   REGION "SELECT WIP BUTTON PULSES"
       "Pop Up: Map Select Button Actuations"(screen_elements := #interface.select_wip_buttons,
                                              actuations_as_ints := #actuations_as_ints);
       #"inst WIP Select Button Pulses"(btns := #actuations_as_ints,
                                        pulses := #actuation_pulses_as_ints);
   END_REGION


   REGION "PERFORM WIP SELECTION"
       "Pop Up: Select WIPs: Perform Selection"(indices := #visable_WIPs_indices,
                                                pulses := #actuation_pulses_as_ints,
                                                visable_WIPs:=#visable_WIPs,
                                                selected_wips_as_bools := #t_selected_WIPs_as_Bools);
   END_REGION


   REGION "MAP SELECTION TO META DATA"
       "Pop Up: Select WIPs: Map to Meta"(actuation_pulses_as_ints := #actuation_pulses_as_ints,
                                          indices := #visable_WIPs_indices,
                                          selected_wips_as_bools := #t_selected_WIPs_as_Bools,
                                          selectable_wips := #meta_data.selectable_wips,
                                          selected_wips := #meta_data.selected_wips);
   END_REGION    


   REGION "HOUSE KEEPING FOR STATION SELECTION CHANGE"
       IF #meta_data.selection_change.selection_change THEN
           "Array.DInt.Fill"(int_in := INT_TO_DINT("NULL_TOKEN"),
                             array_out => #visable_WIPs);
           FOR #i := 0 TO "WIP_COUNT" DO
               #t_selected_WIPs_as_Bools[#i] := FALSE;
           END_FOR;
           "Clear WIP Selection Meta Data"(#meta_data.selected_wips);
       END_IF;
   END_REGION


   REGION "BUILD SELECTABLE WIP LIST"
       IF #meta_data.selection_change.selection_change THEN
           IF "Is_HMI_Station"(#stations.stn[#meta_data.selection_change.station_index]) THEN
               "Pop Up: Select WIPs: Build Selectable List"(saved_WIPs := #saved_WIPs,
                                                            meta_data := #meta_data,
                                                            stations := #stations);
           END_IF;
       END_IF;
   END_REGION


   REGION "SHOW ALL WIPS WHEN FEWER SELECTABLE WIPS THAN BUTTONS"
       IF #meta_data.selection_change.selection_change AND #meta_data.selectable_wips.count - 1 <= "WIP_POPUP_BUTTON_COUNT" THEN
           "Array.DInt.Fill"(int_in := INT_TO_DINT("NULL_TOKEN"),
                             array_out => #visable_WIPs_indices);
           FOR #i := 0 TO #meta_data.selectable_wips.count - 1 DO
               #visable_WIPs[#i] := #meta_data.selectable_wips.wips[#i];
               #visable_WIPs_indices[#i] := #i;
           END_FOR;
       END_IF;
   END_REGION



   REGION "NAVIGATE THROUGH TABLE WHEN MORE SELECTABLE WIPS THAN BUTTONS"
       IF #meta_data.selectable_wips.count - 1 > "WIP_POPUP_BUTTON_COUNT" THEN

           REGION "TABLE NAVIGATION"
               #"inst Table Nav"(first_null_index := #meta_data.selectable_wips.count,
                                 tblData := #meta_data.selectable_wips.wips,
                                 tblDisp := #visable_WIPs,
                                 tableNav := #interface.nav_bar.plc,
                                 rowIndices := #visable_WIPs_indices);
           END_REGION

           REGION "MAP INDICES ON SCANS WHEN SELECTION HASN'T CHANGED"
               IF NOT #meta_data.selection_change.selection_change THEN
                   FOR #i := 0 TO "WIP_POPUP_BUTTON_COUNT" DO
                       #visable_WIPs[#i] := #meta_data.selectable_wips.wips[#visable_WIPs_indices[#i]];
                   END_FOR;
               END_IF;
           END_REGION

           REGION "REMAP INDICES TO TOP WHEN SELECTION HAS CHANGED"
               IF #meta_data.selection_change.selection_change THEN
                   FOR #i := 0 TO "WIP_POPUP_BUTTON_COUNT" DO
                       #visable_WIPs[#i] := INT_TO_DINT(#i);
                       #visable_WIPs_indices[#i] := INT_TO_DINT(#i);
                   END_FOR;
               END_IF;
           END_REGION

       END_IF;
   END_REGION
END_FUNCTION_BLOCK

FUNCTION "Pop Up: Select WIPs: Get Matching WIPs" : Void   // FC125, SCL
{ S7_Optimized_Access := 'TRUE' }
VERSION : 0.1
   VAR_INPUT
      selectable_wips : "Selectable Wips";
      station_wips : "Selectable Wips";
   END_VAR
   VAR_IN_OUT
      matching_wips : "Selectable Wips";
   END_VAR
   VAR_TEMP
      i : Int;
      j : Int;
      t_matching_wips : "Selectable Wips";
   END_VAR
BEGIN
   REGION "COPY TO LOCAL"
       "Array.DInt.Fill"(int_in := INT_TO_DINT("NULL_TOKEN"),
                         array_out => #t_matching_wips.wips);
       #t_matching_wips.count := 0;
   END_REGION

   REGION "COMPARE EACH WIP CODE IN OUTER LIST ..." 
       FOR #i := 0 TO "WIP_COUNT" DO

           REGION "LEAVE LOOP ON FIRST NULL"
               IF #selectable_wips.wips[#i] = "NULL_TOKEN" THEN
                   EXIT;
               END_IF;
           END_REGION

           REGION "WITH EACH IN INNER LIST AND ..."
               FOR #j := 0 TO "WIP_COUNT" DO

                   REGION "LEAVE LOOP ON FIRST NULL"
                       IF #station_wips.wips[#j] = "NULL_TOKEN" THEN
                           EXIT;
                       END_IF;
                   END_REGION

                   REGION "COPY MATCHES"
                       IF #selectable_wips.wips[#i] = #station_wips.wips[#j] THEN
                           #t_matching_wips.wips[#t_matching_wips.count] := #selectable_wips.wips[#i];
                           #t_matching_wips.count += 1;
                       END_IF;
                   END_REGION

               END_FOR;
           END_REGION

       END_FOR;
   END_REGION


   REGION "RETURN"
       #matching_wips := #t_matching_wips;
   END_REGION
END_FUNCTION

FUNCTION "Pop Up: Select WIPs: Build Selectable List" : Void   // FC128, SCL
{ S7_Optimized_Access := 'TRUE' }
VERSION : 0.1
   VAR_INPUT
      stations : "Station: All Stations";
      saved_WIPs : "Recipe: HMI Stations Saved Wips";
   END_VAR
   VAR_IN_OUT
      meta_data : "Setting Meta Data";
   END_VAR
   VAR_TEMP
      wip_index : Int;
      p_outer : Int;
      p_inner : Int;
      t_selectable_WIPs : "Selectable Wips";
      selected_station_WIPs : "Selected Wips";
   END_VAR
BEGIN
   REGION "NO STATIONS SELECTED"
       IF #meta_data.selected_stations.count = 0 THEN
           "Array.DInt.Fill"(int_in := INT_TO_DINT("NULL_TOKEN"),
                             array_out => #t_selectable_WIPs.wips);
           #t_selectable_WIPs.count := 0;
           GOTO RTRN;
       END_IF;
   END_REGION


   REGION "SINGLE STATION SELECTION"
       IF #meta_data.selected_stations.count = 1 THEN
           "Array.DInt.Fill"(int_in := -1,
                             array_out => #t_selectable_WIPs.wips);
           #t_selectable_WIPs.count := 0;
           #wip_index := "WIP.Global_Index_to_HMI_Station_Index"(global_index := "Get First Selected Station"(#meta_data.selected_stations.stns),
                                                                 saved_WIPs := #saved_WIPs);
           "Pop Up: Select WIPs: Map WIP Codes"(wip_station := #saved_WIPs.stn[#wip_index],
                                                selectable_wips := #t_selectable_WIPs);
           GOTO RTRN;
       END_IF;
   END_REGION


   REGION "MULTI STATION SELECTION"

       REGION "CHECK MATCHING: SELECTABLE & NEW STATION"
           #t_selectable_WIPs.wips := #meta_data.selectable_wips.wips;
           "Array.DInt.Fill"(int_in := INT_TO_DINT("NULL_TOKEN"),
                             array_out => #selected_station_WIPs.wips);
           "Map WIP Codes to DInt Array"(station := "WIP.Global_Index_to_Station"(index := #meta_data.selection_change.station_index, wip_stations := #saved_WIPs),
                                         WIP_array := #selected_station_WIPs.wips);
           "Pop Up: Select WIPs: Get Matching WIPs"(selectable_wips := #meta_data.selectable_wips,
                                                    station_wips := #selected_station_WIPs,
                                                    matching_wips := #t_selectable_WIPs);
       END_REGION


   END_REGION


   REGION "RETURN"
   RTRN:
       #meta_data.selectable_wips := #t_selectable_WIPs;
   END_REGION
END_FUNCTION

FUNCTION "Pop Up: Select WIPs: Map WIP Codes" : Void   // FC129, SCL
{ S7_Optimized_Access := 'TRUE' }
VERSION : 0.1
   VAR_INPUT
      wip_station : "WIP: Station";
   END_VAR
   VAR_IN_OUT
      selectable_wips : "Selectable Wips";
   END_VAR
   VAR_TEMP
      i : Int;
      t_selectable_wips : "Selectable Wips";
   END_VAR
BEGIN
   REGION "COPY TO LOCAL"
       #t_selectable_wips := #selectable_wips;
   END_REGION


   REGION "MAP VALUES"
       "Map WIP Codes to DInt Array"(station := #wip_station,
                                     WIP_array := #t_selectable_wips.wips);
   END_REGION


   REGION "COUNT SELECTABLE WIPS"
       #t_selectable_wips.count := "Count Collapsed DInt Array"(null_value := INT_TO_DINT("NULL_TOKEN"),
                                                                array := #t_selectable_wips.wips);
   END_REGION


   REGION "RETURN"
       #selectable_wips := #t_selectable_wips;
   END_REGION
END_FUNCTION

FUNCTION "Pop Up: Select WIPs: Animations" : Void   // FC134, SCL
{ S7_Optimized_Access := 'TRUE' }
VERSION : 0.1
   VAR_INPUT
      selectable_WIP_count : Int;
      selected_WIPs : Array[0.."WIP_COUNT"] of Bool;
      visable_WIPs : Array[0.."WIP_POPUP_BUTTON_COUNT"] of DInt;
      visable_WIPs_indices : Array[0.."WIP_POPUP_BUTTON_COUNT"] of Int;
      wip_library : "Recipe: Wip Text Library";
   END_VAR
   VAR_IN_OUT
      interface : "Select WIP";
   END_VAR
   VAR_TEMP
      i : Int;
      labels : Array[0.."WIP_POPUP_BUTTON_COUNT"] of String;
      t_interface : "Select WIP";
      t_selected_WIPs : Array[0.."WIP_COUNT"] of Int;
      visable_WIP_count : Int;
   END_VAR
BEGIN
   REGION "COPY TO LOCAL"
       #t_interface := #interface;
   END_REGION


   REGION "ANIMATE CLOSE SCREEN BUTTON"
       #t_interface.close_screen.animate := "Bool.Animate"(true_color := "GREEN_LIGHT_BACKGROUND",
                                                           false_color := "RED_LIGHT_BACKGROUND",
                                                           evaluation_signal := #t_interface.close_screen.actuate);
   END_REGION


   REGION "ANIMATE WIP SELECT BUTTONS" 

       REGION "WIP LABELS"
           FOR #i := 0 TO "WIP_POPUP_BUTTON_COUNT" DO
               #labels[#i] := WSTRING_TO_STRING("WIP.Code_to_WString"(wipTxtLib := #wip_library, code := #visable_WIPs[#i]));
           END_FOR;
       END_REGION

       REGION "CONVERT BOOLS TO INT FOR MOVE BLOCK VARIANT"
           FOR #i := 0 TO "WIP_COUNT" DO
               #t_selected_WIPs[#i].%X0 := #selected_WIPs[#i];
           END_FOR;
       END_REGION

       REGION "ANIMATE"
           #visable_WIP_count := "Count Collapsed DInt Array"(null_value := INT_TO_DINT("NULL_TOKEN"),
                                                              array := #visable_WIPs);
           "Animate Array: PB Data"(labels := #labels,
                                    pb_data := #t_interface.select_wip_buttons,
                                    selected_elements := #t_selected_WIPs,
                                    visible_elements := #visable_WIPs_indices,
                                    visible_pb_count := #visable_WIP_count);
       END_REGION

   END_REGION


   REGION "NAV BAR"
       "Pop Up: Nav Bar: Animate"(selectable_element_count := #selectable_WIP_count - 1,
                                  visible_rows := "WIP_POPUP_BUTTON_COUNT",
                                  nav_bar := #t_interface.nav_bar);
   END_REGION


   REGION "DRAW"
       #interface := #t_interface;
   END_REGION
END_FUNCTION

FUNCTION "Pop Up: Select WIPs: Perform Selection" : Void   // FC137, SCL
{ S7_Optimized_Access := 'TRUE' }
VERSION : 0.1
   VAR_INPUT
      indices : Array[0.."WIP_POPUP_BUTTON_COUNT"] of DInt;
      pulses : Array[0.."WIP_POPUP_BUTTON_COUNT"] of Int;
      visable_WIPs : Array[0.."WIP_POPUP_BUTTON_COUNT"] of DInt;
   END_VAR
   VAR_IN_OUT
      selected_wips_as_bools : Array[0.."WIP_COUNT"] of Bool;
   END_VAR
   VAR_TEMP
      i : Int;
      t_selected_wips_as_bools : Array[0.."WIP_COUNT"] of Bool;
   END_VAR
BEGIN
   REGION "NOTES"
       (*
           The same wip code can exist in several hmi stations, so 
           selected wips are stored by generating an array of codes.
           Later, the codes can be checked at each station for station 
           modificatins.
           This function starts the process by checking the visable indices
           array (a list of pointers to rows in the selectable wip array).
           If an actuation occurs on a button, visible[x] will give the row 
           number of the wip code in the selectable wip array.
           The row number in the selected wip array is then set to true.
           The toggeled state together with the pulse allows the selected 
           wips list to be rebuilt easily.
       *)
   END_REGION


   REGION "COPY TO LOCAL"
       #t_selected_wips_as_bools := #selected_wips_as_bools;
   END_REGION


   REGION "CHECK INDEX ARRAY"
       FOR #i := 0 TO "WIP_POPUP_BUTTON_COUNT" DO

           REGION "EXIT ON NULL"
               IF #visable_WIPs[#i] = "NULL_TOKEN" THEN
                   EXIT;
               END_IF;
           END_REGION

           REGION "TOGGLE WIP SELECT STATE"
               "Toggle"(pulse := #pulses[#i].%X0,
                        state := #t_selected_wips_as_bools[DINT_TO_INT(#indices[#i])]);
           END_REGION

       END_FOR;
   END_REGION


   REGION "RETURN"
       #selected_wips_as_bools := #t_selected_wips_as_bools;
   END_REGION
END_FUNCTION

FUNCTION "Pop Up: Select WIPs: Map to Meta" : Void   // FC138, SCL
{ S7_Optimized_Access := 'TRUE' }
VERSION : 0.1
   VAR_INPUT
      actuation_pulses_as_ints : Array[0.."WIP_POPUP_BUTTON_COUNT"] of Int;
      indices : Array[0.."WIP_POPUP_BUTTON_COUNT"] of DInt;
      selected_wips_as_bools : Array[0.."WIP_COUNT"] of Bool;
      selectable_wips : "Selectable Wips";
   END_VAR
   VAR_IN_OUT
      selected_wips : "Selected Wips";
   END_VAR
   VAR_TEMP
      rebuild_selected_wips : Bool;
      i : Int;
      t_selected_wips : "Selected Wips";
   END_VAR
BEGIN
   REGION "NOTES"
       (*
           This function has two states.
           The first state checks for any selection pulse.
           On such a pulse, the selected wip code array is filled
           with nulls, the selected wip counter is reset, and the 
           state flag to rebuild the array is set.
           In the rebuild array state, each element of the selected
           wip array of bools is checked. 
           If true, the code from the corresponding selectable wip
           code array is saved to the selected wip code array and 
           the selected wip count is incremented.
           When this function has completed, the array of selected wips
           in meta data section of the hmi settings db will be up to 
           date.
          *)
   END_REGION


   REGION "COPY TO LOCAL"
       #t_selected_wips := #selected_wips;
   END_REGION


   REGION "SCAN FOR PULSES, INITIALIZE AND SET STATE"
       FOR #i := 0 TO "WIP_POPUP_BUTTON_COUNT" DO
           IF #actuation_pulses_as_ints[#i].%X0 THEN
               "Array.DInt.Fill"(int_in := INT_TO_DINT("NULL_TOKEN"),
                                 array_out => #t_selected_wips.wips);
               #t_selected_wips.count := 0;
               #rebuild_selected_wips := TRUE;
               EXIT;
           END_IF;
       END_FOR;
   END_REGION


   REGION "REBUILD ARRAY, INCREMENT SELECTED WIP COUNT"
       IF #rebuild_selected_wips THEN
           FOR #i := 0 TO "WIP_COUNT" DO
               IF #selected_wips_as_bools[#i] THEN
                   #t_selected_wips.wips[#t_selected_wips.count] := #selectable_wips.wips[#i];
                   #t_selected_wips.count += 1;
               END_IF;
           END_FOR;
       END_IF;
   END_REGION


   REGION "RETURN"
       #selected_wips := #t_selected_wips;
   END_REGION
END_FUNCTION

// folder: HMI: Warehouse/RSP Simulation

FUNCTION_BLOCK "Sim: from Global"   // FB26, SCL
{ S7_Optimized_Access := 'TRUE' }
VERSION : 0.1
   VAR_INPUT
      stns : "Station: All Stations";
   END_VAR
   VAR_IN_OUT
      simStations : "Simulated Stations";
   END_VAR
   VAR
      old : Struct
         nextGrp : Bool;
         prevGrp : Bool;
      END_STRUCT;
   END_VAR
   VAR_TEMP
      animate : USInt;
      btnCount : Int;
      currentBtn : Bool;
      dzLabel : WString;
      firstStn : Int;
      i : Int;
      intBox : Int;
      j : Int;
      kp8Color : DWord;
      label : WString;
      oldBtn : Bool;
      pSim : Int;
      pStn : Int;
   END_VAR
   VAR CONSTANT
      space : WString := WSTRING#' ';
      lead0 : WString := WSTRING#'0';
      volvo16 : WString := WSTRING#'VOLVO 16';
   END_VAR
BEGIN
   REGION "COPY TO LOCAL"
       #firstStn := #simStations.firstStn;
   END_REGION

   REGION "RESOLVE STATION POINTER"

       REGION "PROCESS NEXT GROUP PRESS"

           REGION "COPY TO LOCAL"
               #currentBtn := #simStations.down.actuate;
               #oldBtn := #old.nextGrp;
           END_REGION

           REGION "FALLING EDGE OF NEXT GROUP"
               IF NOT #currentBtn AND #oldBtn THEN

                   REGION "INCREMENT FIRST STATION"
                       #firstStn += "simKP8Count";
                   END_REGION

                   REGION "UPPER LIMIT ROLL OVER"
                       IF #firstStn > "STATION_COUNT" THEN
                           #firstStn -= "STATION_COUNT" + 1;
                       END_IF;
                   END_REGION

               END_IF;
           END_REGION

           REGION "NEXT GROUP CHANGE DETECTION"
               #old.nextGrp := #currentBtn;
           END_REGION

       END_REGION

       REGION "PROCESS PREVIOUS GROUP PRESS"

           REGION "COPY TO LOCAL"
               #currentBtn := #simStations.up.actuate;
               #oldBtn := #old.prevGrp;
           END_REGION

           REGION "FALLING EDGE OF PREVIOUS GROUP"
               IF NOT #currentBtn AND #oldBtn THEN

                   REGION "DECREMENT FIRST STATION"
                       #firstStn -= "simKP8Count";
                   END_REGION

                   REGION "LOWER LIMIT ROLL OVER"
                       IF #firstStn < 0 THEN
                           #firstStn += "STATION_COUNT" + 1;
                       END_IF;
                   END_REGION

               END_IF;
           END_REGION

           REGION "PREVIOUS GROUP CHANGE DETECTION"
               #old.prevGrp := #currentBtn;
           END_REGION

       END_REGION

   END_REGION

   REGION "FOR EACH BUTTON"
       FOR #i := 0 TO 11 DO

           REGION "CALCULATE POINTER"
               #pStn := #i + #firstStn;
               #pSim := #i;
           END_REGION

           REGION "UPPER LIMIT ROLL OVER"
               IF #pStn > "STATION_COUNT" THEN
                   #pStn := #firstStn + #i - "STATION_COUNT" - 1;
               END_IF;
           END_REGION

           REGION "COPY TO LOCAL"
               #kp8Color := #stns.stn[#pStn].wipCmpts.ioData.kp8.tempOut;
           END_REGION

           REGION "LABEL STATIONS"

               REGION "DETERMINE LINE LABEL"
                   #label := #stns.stn[#pStn].id.lineName;
                   IF #label = #volvo16 THEN
                       #label := WSTRING#'V16';
                   END_IF;
               END_REGION

               REGION "DETERMINE DROP ZONE LABEL"
                   #intBox := USINT_TO_INT(#stns.stn[#pStn].id.dropZone);
                   IF #intBox <= 9 THEN
                       #dzLabel := CONCAT_WSTRING(IN1 := #lead0,
                                                  IN2 := "Strip Sign"(INT_TO_WSTRING(#intBox)));
                   END_IF;
                   IF #intBox >= 10 THEN
                       #dzLabel := "Strip Sign"(INT_TO_WSTRING(#intBox));
                   END_IF;
               END_REGION

               REGION "WRITE LABEL"
                   #label := CONCAT_WSTRING(IN1 := #label,
                                            IN2 := #space,
                                            IN3 := #dzLabel);
                   #simStations.me[#pSim].stn.label := #label;
               END_REGION

           END_REGION

           REGION "ANIMATE STATION LABEL"
               #simStations.me[#pSim].stn.animate := "GRAY_BACKGROUND";
           END_REGION

           REGION "FOR EACH BUTTON"
               FOR #j := 0 TO "STATION_BUTTON_COUNT" DO

                   REGION "COLOR BUTTONS"
                       #animate := "KP8 Driver: HMI Emulator: Animation"(kp8Color := #kp8Color,
                                                                btnNumber := #j);
                       #simStations.me[#pSim].btn.animate[#j] := #animate;
                   END_REGION

                   REGION "WRITE BUTTON LABELS"
                       #intBox := "Pointer Calc: KP8 Labels"(#j);
                       #label := "Strip Sign"(INT_TO_WSTRING(#intBox));
                       #simStations.me[#pSim].btn.labels[#j] := #label;
                   END_REGION

               END_FOR;
           END_REGION

       END_FOR;
   END_REGION

   REGION "SAVE FIRST STATION"
       #simStations.firstStn := #firstStn;
   END_REGION

   REGION "ANIMATE NEXT GROUP PRESS"
       #simStations.down.animate := "Bool.Animate"(true_color := "GREEN_LIGHT_BACKGROUND",
                                                   false_color := "GRAY_BACKGROUND",
                                                   evaluation_signal := #simStations.down.actuate);
   END_REGION

   REGION "ANIMATE PREV GROUP PARESS"
       #simStations.up.animate := "Bool.Animate"(true_color := "GREEN_LIGHT_BACKGROUND",
                                                 false_color := "GRAY_BACKGROUND",
                                                 evaluation_signal := #simStations.up.actuate);
   END_REGION
END_FUNCTION_BLOCK

FUNCTION "Sim: to Global" : Void   // FC23, SCL
{ S7_Optimized_Access := 'TRUE' }
VERSION : 0.1
   VAR_INPUT
      simStns : "Simulated Stations";
   END_VAR
   VAR_IN_OUT
      stations : "Station: All Stations";
   END_VAR
   VAR_TEMP
      i : Int;
      j : Int;
      pSim : Int;
      pStn : Int;
   END_VAR
BEGIN
   REGION "COPY TO LOCAL"
       // #btnCount := "btnCount";
       // #firstStn := #simStns.firstStn;
       // #simKP8Count := "simKP8Count";
       // #stnCount := "stnCount";
   END_REGION

   REGION "FOR EACH STATION"
       FOR #i := 0 TO "simKP8Count" DO

           REGION "CALCULATE POINTER"
               #pStn := #i + #simStns.firstStn;
               #pSim := #i;
           END_REGION

           REGION "UPPER LIMIT ROLL OVER"
               IF #pStn > "STATION_COUNT" THEN
                   #pStn := #simStns.firstStn + #i - "STATION_COUNT" - 1;
               END_IF;
           END_REGION

           REGION "COPY SIMULATED PRESSES"
               #stations.stn[#pStn].wipCmpts.ioData.kp8.input.%B1 := #simStns.me[#pSim].btn.actuate;
           END_REGION

       END_FOR;
   END_REGION
END_FUNCTION

FUNCTION "Sim: KP8 Animations" : Word   // FC84, SCL
{ S7_Optimized_Access := 'TRUE' }
VERSION : 0.1
   VAR_INPUT
      pbs : DWord;
   END_VAR
   VAR_TEMP
      ret : Word;
   END_VAR
BEGIN
   #"Sim: KP8 Animations".%B1 := #pbs.%B0;
   #"Sim: KP8 Animations".%B0 := #pbs.%B1;
END_FUNCTION

// folder: Linked List

FUNCTION_BLOCK "Linked List"   // FB29, SCL
{ S7_Optimized_Access := 'TRUE' }
VERSION : 0.1
   VAR_IN_OUT
      interface : "Linked List: Method Interface";
   END_VAR
   VAR
      list : "Linked List: List";
   END_VAR
   VAR CONSTANT
      TERMINAL_BEHAVIOR : String := 'open';
   END_VAR
BEGIN
   REGION "APPEND"
       IF #interface.append.in.request THEN
           "Linked List: Append"(terminal_behavior := #TERMINAL_BEHAVIOR,
                                 commands := #interface.append,
                                 list := #list);
       END_IF;
   END_REGION

   REGION "DELETE"
       IF #interface.delete.in.request THEN
           "Linked List: Delete"(commands := #interface.delete,
                                 list := #list);
       END_IF;
   END_REGION

   REGION "DISPLAY"
       IF #interface.display.in.request THEN
           "Linked List: Display"(commands := #interface.display,
                                  list := #list);
       END_IF;
   END_REGION

   REGION "INSERT"
       IF #interface.insert.in.request THEN
           "Linked List: Insert"(terminal_behavior := #TERMINAL_BEHAVIOR,
                                 commands := #interface.insert,
                                 list := #list);
       END_IF;
   END_REGION

   REGION "RESET"
       IF #interface.reset.in.request THEN
           "Linked List: Reset"(commands := #interface.reset,
                                list := #list);
       END_IF;
   END_REGION

   REGION "REVERSE"
       IF #interface.reverse.in.request THEN
           "Linked List: Reverse"(commands := #interface.reverse,
                                  list := #list);
       END_IF;
   END_REGION

   REGION "SEARCH"
       IF #interface.search.in.request THEN
           "Linked List: Search"(commands := #interface.search,
                                 list := #list);
       END_IF;
   END_REGION
END_FUNCTION_BLOCK

FUNCTION "Linked List: Private: Clear Node" : Void   // FC156, SCL
{ S7_Optimized_Access := 'TRUE' }
VERSION : 0.1
   VAR_IN_OUT
      node : "Linked List: Node";
   END_VAR
   VAR_TEMP
      ret : "Linked List: Node";
   END_VAR
BEGIN
   #ret.meta.key := "NULL_TOKEN";
   #ret.meta.next := "NULL_TOKEN";
   #node := #ret;
END_FUNCTION

FUNCTION "Linked List: Private: Get Head" : "Linked List: Node"   // FC157, SCL
{ S7_Optimized_Access := 'TRUE' }
VERSION : 0.1
   VAR_INPUT
      list : "Linked List: List";
   END_VAR
   VAR_TEMP
      pointer_list : DInt;
      ret : "Linked List: Node";
   END_VAR
BEGIN
   FOR #pointer_list := 0 TO "LINKED_LIST_LENGTH" DO
       IF #list.me[#pointer_list].meta.is_head THEN
           #ret := #list.me[#pointer_list];
           EXIT;
       END_IF;
   END_FOR;
   #"Linked List: Private: Get Head" := #ret;
END_FUNCTION

FUNCTION "Linked List: Private: Before" : Void   // FC158, SCL
{ S7_Optimized_Access := 'TRUE' }
VERSION : 0.1
   VAR_IN_OUT
      next_node : "Linked List: Node";   // next_node goes after node
      node : "Linked List: Node";   // node goes before next_node
   END_VAR
BEGIN
   #node.meta.next := #next_node.meta.key;
   IF #next_node.meta.is_head THEN
       #next_node.meta.is_head := FALSE;
       #node.meta.is_head := TRUE;
   END_IF;
END_FUNCTION

FUNCTION "Linked List: Private: Tail Swap" : Void   // FC159, SCL
{ S7_Optimized_Access := 'TRUE' }
VERSION : 0.1
   VAR_IN_OUT
      new_tail : "Linked List: Node";
      old_tail : "Linked List: Node";
   END_VAR
BEGIN
   #new_tail.meta.is_tail := TRUE;
   #old_tail.meta.is_tail := FALSE;
END_FUNCTION

FUNCTION "Linked List: Private: Head Swap" : Void   // FC160, SCL
{ S7_Optimized_Access := 'TRUE' }
VERSION : 0.1
   VAR_IN_OUT
      new_head : "Linked List: Node";
      old_head : "Linked List: Node";
   END_VAR
BEGIN
   #new_head.meta.is_head := TRUE;
   #old_head.meta.is_head := FALSE;
END_FUNCTION

FUNCTION "Linked List: Private: Get Next" : "Linked List: Node"   // FC161, SCL
{ S7_Optimized_Access := 'TRUE' }
VERSION : 0.1
   VAR_INPUT
      current : "Linked List: Node";
      list : "Linked List: List";
   END_VAR
   VAR_TEMP
      ret : "Linked List: Node";
   END_VAR
BEGIN
   "Linked List: Private: Clear Node"(#ret);
   IF #list.me[#current.meta.key].meta.next <> "NULL_TOKEN" THEN
       #ret := #list.me[#current.meta.next];
   END_IF;
   #"Linked List: Private: Get Next" := #ret;
END_FUNCTION

FUNCTION "Linked List: Private: Get Previous" : "Linked List: Node"   // FC162, SCL
{ S7_Optimized_Access := 'TRUE' }
VERSION : 0.1
   VAR_INPUT
      current : "Linked List: Node";
      list : "Linked List: List";
   END_VAR
   VAR_TEMP
      list_pointer : DInt;
      ret : "Linked List: Node";
   END_VAR
BEGIN
   "Linked List: Private: Clear Node"(#ret);
   FOR #list_pointer := 0 TO "LINKED_LIST_LENGTH" DO
       IF #list.me[#list_pointer].meta.next = #current.meta.key THEN
           #ret := #list.me[#list_pointer];
           EXIT;
       END_IF;
   END_FOR;
   #"Linked List: Private: Get Previous" := #ret;
END_FUNCTION

FUNCTION "Linked List: Private: After" : Void   // FC163, SCL
{ S7_Optimized_Access := 'TRUE' }
VERSION : 0.1
   VAR_IN_OUT
      node : "Linked List: Node";
      previous_node : "Linked List: Node";
   END_VAR
BEGIN
   #node.meta.next := #previous_node.meta.next;
   #previous_node.meta.next := #node.meta.key;
   IF #previous_node.meta.is_tail THEN
       #previous_node.meta.is_tail := FALSE;
       #node.meta.is_tail := TRUE;
   END_IF;
END_FUNCTION

FUNCTION "Linked List: Private: Head an Empty List" : Void   // FC164, SCL
{ S7_Optimized_Access := 'TRUE' }
VERSION : 0.1
   VAR_INPUT
      data : "Linked List: Node: Data";
      terminal_behavior : String;   // 'open': head's previous and tail's next are null nodes; 'closed': head's previous is tail, tail's next is head
   END_VAR
   VAR_IN_OUT
      list : "Linked List: List";
   END_VAR
BEGIN
   #list.me[0].data := #data;
   #list.me[0].meta.key := 0;
   IF #terminal_behavior = 'open' THEN
       #list.me[0].meta.next := "NULL_TOKEN";
   END_IF;
   IF #terminal_behavior = 'closed' THEN
       #list.me[0].meta.next := 0;
   END_IF;
   #list.me[0].meta.is_head := TRUE;
   #list.me[0].meta.is_tail := TRUE;
END_FUNCTION

FUNCTION "Linked List: Private: Is Empty" : Bool   // FC165, SCL
{ S7_Optimized_Access := 'TRUE' }
VERSION : 0.1
   VAR_INPUT
      list : "Linked List: List";
   END_VAR
   VAR_TEMP
      pointer_list : DInt;
      ret : Bool;
   END_VAR
BEGIN
   #ret := TRUE;
   FOR #pointer_list := 0 TO "LINKED_LIST_LENGTH" DO
       IF #list.me[#pointer_list].meta.key <> "NULL_TOKEN" THEN
           #ret := FALSE;
           EXIT;
       END_IF;
   END_FOR;
   #"Linked List: Private: Is Empty" := #ret;
END_FUNCTION

FUNCTION "Linked List: Private: Get Tail" : "Linked List: Node"   // FC166, SCL
{ S7_Optimized_Access := 'TRUE' }
VERSION : 0.1
   VAR_IN_OUT
      list : "Linked List: List";
   END_VAR
   VAR_TEMP
      pointer_list : Int;
      next_node : UInt;
      ret : "Linked List: Node";
   END_VAR
BEGIN
   FOR #pointer_list := 0 TO "LINKED_LIST_LENGTH" DO
       IF #list.me[#pointer_list].meta.is_tail THEN
           #ret := #list.me[#pointer_list];
           EXIT;
       END_IF;
   END_FOR;
   #"Linked List: Private: Get Tail" := #ret;
END_FUNCTION

FUNCTION "Linked List: Private: Is Full" : Bool   // FC167, SCL
{ S7_Optimized_Access := 'TRUE' }
VERSION : 0.1
   VAR_INPUT
      list : "Linked List: List";
   END_VAR
   VAR_TEMP
      pointer_list : DInt;
      ret : Bool;
   END_VAR
BEGIN
   #ret := TRUE;
   FOR #pointer_list := 0 TO "LINKED_LIST_LENGTH" DO
       IF #list.me[#pointer_list].meta.key = "NULL_TOKEN" THEN
           #ret := FALSE;
           EXIT;
       END_IF;
   END_FOR;
   #"Linked List: Private: Is Full" := #ret;
END_FUNCTION

FUNCTION "Linked List: Private: Next Empty Node" : DInt   // FC168, SCL
{ S7_Optimized_Access := 'TRUE' }
VERSION : 0.1
   VAR_IN_OUT
      list : "Linked List: List";
   END_VAR
   VAR_TEMP
      node : "Linked List: Node";
      pointer_list : Int;
      ret : DInt;
   END_VAR
BEGIN
   #ret := "NULL_TOKEN";
   FOR #pointer_list := 0 TO "LINKED_LIST_LENGTH" DO
       IF #list.me[#pointer_list].meta.key = "NULL_TOKEN" THEN
           #ret := INT_TO_DINT(#pointer_list);
           EXIT;
       END_IF;
   END_FOR;
   #"Linked List: Private: Next Empty Node" := #ret;
END_FUNCTION

FUNCTION "Linked List: Append" : Void   // FC169, SCL
{ S7_Optimized_Access := 'TRUE' }
VERSION : 0.1
   VAR_INPUT
      terminal_behavior : String;
   END_VAR
   VAR_IN_OUT
      commands : "Linked List: Method Interface: Append";
      list : "Linked List: List";
   END_VAR
   VAR_TEMP
      clear_commands : "Linked List: Method Interface: Append";
      head : "Linked List: Node";
      pointer_new_node : DInt;
      tail : "Linked List: Node";
   END_VAR
   VAR CONSTANT
      no_error : String := 'no error';
      list_full : String := 'appended to full list';
      no_tail_found : String := 'no tail found while trying to append';
      appended_as_head : String := 'appended as head of list';
   END_VAR
BEGIN
   REGION "NOTES"
       (*
       Append adds a node to the end of the list.
       Last edit: 2021-10-05
       *)
   END_REGION

   REGION "APPEND TO FULL LIST"
       IF "Linked List: Private: Is Full"(#list) THEN
           #commands := #clear_commands;
           #commands.out.error := TRUE;
           #commands.out.error_message := #list_full;
           RETURN;
       END_IF;
   END_REGION

   REGION "APPEND TO EMPTY LIST"
       IF "Linked List: Private: Is Empty"(#list) THEN
           "Linked List: Private: Head an Empty List"(data := #commands.in.data,
                                                      terminal_behavior := #terminal_behavior,
                                                      list := #list);
           #commands := #clear_commands;
           #commands.out.done := TRUE;
           #commands.out.error_message := #appended_as_head;
           RETURN;
       END_IF;
   END_REGION

   REGION "FIND TAIL"
       #tail := "Linked List: Private: Get Tail"(#list);
   END_REGION

   REGION "EXIT CONDITION: TAIL NOT FOUND"
       IF #tail.meta.key = "NULL_TOKEN" THEN
           #commands := #clear_commands;
           #commands.out.error := TRUE;
           #commands.out.error_message := #no_tail_found;
           RETURN;
       END_IF;
   END_REGION

   REGION "FIND FIRST NULL"
       #pointer_new_node := "Linked List: Private: Next Empty Node"(#list);
   END_REGION

   REGION "APPENDED NODE IS AFTER TAIL"
       #list.me[#pointer_new_node].data := #commands.in.data;
       #list.me[#pointer_new_node].meta.key := #pointer_new_node;
       "Linked List: Private: After"(node := #list.me[#pointer_new_node],
                                     previous_node := #list.me[#tail.meta.key]);
   END_REGION

   REGION "EXIT CONDITION: SUCCESS"
       #commands := #clear_commands;
       #commands.out.done := TRUE;
       #commands.out.error_message := #no_error;
   END_REGION
END_FUNCTION

FUNCTION "Linked List: Delete" : Void   // FC170, SCL
{ S7_Optimized_Access := 'TRUE' }
VERSION : 0.1
   VAR_IN_OUT
      commands : "Linked List: Method Interface: Delete";
      list : "Linked List: List";
   END_VAR
   VAR_TEMP
      blank_node : "Linked List: Node";
      clear_commands : "Linked List: Method Interface: Delete";
      current : "Linked List: Node";
      found : Bool;
      next : "Linked List: Node";
      pointer_list : DInt;
      previous : "Linked List: Node";
      search_commands : "Linked List: Method Interface: Search";
   END_VAR
   VAR CONSTANT
      no_error : String := 'no error';
      delete_from_empty : String := 'deleted from an empty list.';
   END_VAR
BEGIN
   REGION "EXIT CONDITION: LIST IS EMPTY"
       IF "Linked List: Private: Is Empty"(#list) THEN
           #commands := #clear_commands;
           #commands.out.error := TRUE;
           #commands.out.error_message := #delete_from_empty;
       END_IF;
   END_REGION

   REGION "DELETE"
       #current := #commands.in.node;
       #previous := "Linked List: Private: Get Previous"(current := #current,
                                                         list := #list);
       #next := "Linked List: Private: Get Next"(current := #current,
                                                 list := #list);
       IF #current.meta.is_head AND NOT #current.meta.is_tail THEN
           "Linked List: Private: Head Swap"(new_head := #list.me[#next.meta.key],
                                             old_head := #list.me[#current.meta.key]);
       END_IF;
       IF NOT #current.meta.is_head AND #current.meta.is_tail THEN
           "Linked List: Private: Tail Swap"(new_tail := #list.me[#previous.meta.key],
                                             old_tail := #list.me[#current.meta.key]);
       END_IF;
       IF NOT #current.meta.is_head THEN
           #list.me[#previous.meta.key].meta.next := #next.meta.key;
       END_IF;
       "Linked List: Private: Clear Node"(#list.me[#current.meta.key]);
   END_REGION

   REGION "COMMANDS OUT"
       #commands := #clear_commands;
       #commands.out.done := TRUE;
       #commands.out.error_message := #no_error;
   END_REGION
END_FUNCTION

FUNCTION "Linked List: Search" : Void   // FC171, SCL
{ S7_Optimized_Access := 'TRUE' }
VERSION : 0.1
   VAR_IN_OUT
      commands : "Linked List: Method Interface: Search";
      list : "Linked List: List";
   END_VAR
   VAR_TEMP
      clear_commands : "Linked List: Method Interface: Search";
      found : Bool;
      pointer_list : DInt;
   END_VAR
   VAR CONSTANT
      no_error : String := 'no error';
      searched_empty_list : String := 'searched empty list';
   END_VAR
BEGIN
   REGION "EXIT CONDITION: SEARCHED EMPTY LIST"
       IF "Linked List: Private: Is Empty"(#list) THEN
           #commands := #clear_commands;
           #commands.out.not_found := TRUE;
           #commands.out.error := TRUE;
           #commands.out.error_message := #searched_empty_list;
           RETURN;
       END_IF;
   END_REGION

   REGION "SEARCH"
       FOR #pointer_list := 0 TO "LINKED_LIST_LENGTH" DO
           IF #list.me[#pointer_list].data = #commands.in.data THEN
               #found := TRUE;
               EXIT;
           END_IF;
       END_FOR;
   END_REGION

   REGION "FOUND"
       IF #found THEN
           #commands := #clear_commands;
           #commands.out.done := TRUE;
           #commands.out.found := TRUE;
           #commands.out.returned_node := #list.me[#pointer_list];
           #commands.out.error_message := #no_error;
           RETURN;
       END_IF;
   END_REGION

   REGION "NOT FOUND"
       IF NOT #found THEN
           #commands := #clear_commands;
           #commands.out.done := TRUE;
           #commands.out.not_found := TRUE;
           RETURN;
       END_IF;
   END_REGION
END_FUNCTION

FUNCTION "Linked List: Display" : Void   // FC172, SCL
{ S7_Optimized_Access := 'TRUE' }
VERSION : 0.1
   VAR_IN_OUT
      commands : "Linked List: Method Interface: Display";
      list : "Linked List: List";
   END_VAR
   VAR_TEMP
      clear_commands : "Linked List: Method Interface: Display";
   END_VAR
BEGIN
   #commands := #clear_commands;
   #commands.out.list := #list;
   #commands.out.done := TRUE;
END_FUNCTION

FUNCTION "Linked List: Insert" : Void   // FC173, SCL
{ S7_Optimized_Access := 'TRUE' }
VERSION : 0.1
   VAR_INPUT
      terminal_behavior : String;
   END_VAR
   VAR_IN_OUT
      commands : "Linked List: Method Interface: Insert";
      list : "Linked List: List";
   END_VAR
   VAR_TEMP
      clear_commands : "Linked List: Method Interface: Insert";
      current : "Linked List: Node";
      next_empty_node_index : DInt;
      previous : "Linked List: Node";
      next : "Linked List: Node";
   END_VAR
   VAR CONSTANT
      no_error : String := 'no error';
      inserted_into_full : String := 'attempted to insert into full list. delete a node and try again.';
      appended_as_head : String := 'appended as head of list';
   END_VAR
BEGIN
   REGION "EXIT CONDITION: INSERTED INTO FULL LIST"
       IF "Linked List: Private: Is Full"(#list) THEN
           #commands := #clear_commands;
           #commands.out.error := TRUE;
           #commands.out.error_message := #inserted_into_full;
           RETURN;
       END_IF;
   END_REGION

   REGION "EXIT CONDITION: INSERTED INTO EMPTY LIST"
       IF "Linked List: Private: Is Empty"(#list) THEN
           "Linked List: Private: Head an Empty List"(data := #commands.in.data,
                                                      terminal_behavior := #terminal_behavior,
                                                      list := #list);
           #commands := #clear_commands;
           #commands.out.error := TRUE;
           #commands.out.error_message := #appended_as_head;
           RETURN;
       END_IF;
   END_REGION

   REGION "GET INDEX OF NEXT EMPTY NODE"
       #next_empty_node_index := "Linked List: Private: Next Empty Node"(#list);
   END_REGION

   REGION "PREVIOUS, CURRENT, AND NEXT NODES"
       #current := #commands.in.target_node;
       #previous := "Linked List: Private: Get Previous"(current := #current,
                                                         list := #list);
       #next := #current;
   END_REGION

   REGION "INSERT BEFORE TARGET NODE"
       // new node's data becomes command data
       #list.me[#next_empty_node_index].data := #commands.in.data;
       // new node's key becomes array index
       #list.me[#next_empty_node_index].meta.key := #next_empty_node_index;
       // shorten name for indexing
       #current := #list.me[#next_empty_node_index];
       // insert
       IF NOT #next.meta.is_head THEN
           "Linked List: Private: After"(node := #list.me[#current.meta.key],
                                         previous_node := #list.me[#previous.meta.key]);
       END_IF;
       "Linked List: Private: Before"(next_node := #list.me[#next.meta.key],
                                      node := #list.me[#current.meta.key]);
   END_REGION

   REGION "COMMANDS OUT"
       #commands := #clear_commands;
       #commands.out.done := TRUE;
       #commands.out.error_message := #no_error;
   END_REGION
END_FUNCTION

FUNCTION "Linked List: Reverse" : Void   // FC174, SCL
{ S7_Optimized_Access := 'TRUE' }
VERSION : 0.1
   VAR_IN_OUT
      commands : "Linked List: Method Interface: Reverse";
      list : "Linked List: List";
   END_VAR
   VAR_TEMP
      clear_commands : "Linked List: Method Interface: Reverse";
      current : "Linked List: Node";
      next : "Linked List: Node";
      previous : "Linked List: Node";
      null_node : "Linked List: Node";
   END_VAR
   VAR CONSTANT
      no_error : String := 'no error';
      reversed_empty_list : String := 'reversed empty list';
   END_VAR
BEGIN
   IF "Linked List: Private: Is Empty"(#list) THEN
       #commands := #clear_commands;
       #commands.out.error := TRUE;
       #commands.out.error_message := #reversed_empty_list;
       RETURN;
   END_IF;

   "Linked List: Private: Clear Node"(#null_node);
   #previous := #null_node;
   #current := "Linked List: Private: Get Head"(#list);
   #list.me[#current.meta.key].meta.is_head := FALSE;
   #list.me[#current.meta.key].meta.is_tail := TRUE;
   WHILE #current.meta.next <> "NULL_TOKEN" DO
       #next := #list.me[#current.meta.next];
       #list.me[#current.meta.key].meta.next := #previous.meta.key;
       #previous := #current;
       #current := #next;
       #list.me[#current.meta.key].meta.is_head := FALSE;
       #list.me[#current.meta.key].meta.is_tail := FALSE;
   END_WHILE;
   #list.me[#current.meta.key].meta.next := #previous.meta.key;
   #list.me[#current.meta.key].meta.is_head := TRUE;
   #list.me[#current.meta.key].meta.is_tail := FALSE;

   #commands := #clear_commands;
   #commands.out.done := TRUE;
   #commands.out.error_message := #no_error;
END_FUNCTION

FUNCTION "Linked List: Reset" : Void   // FC175, SCL
{ S7_Optimized_Access := 'TRUE' }
VERSION : 0.1
   VAR_IN_OUT
      commands : "Linked List: Method Interface: Reset";
      list : "Linked List: List";
   END_VAR
   VAR_TEMP
      blank_node : "Linked List: Node";
      list_pointer : DInt;
      clear_commands : "Linked List: Method Interface: Reset";
   END_VAR
BEGIN
   FOR #list_pointer := 0 TO "LINKED_LIST_LENGTH" DO
       "Linked List: Private: Clear Node"(#list.me[#list_pointer]);
   END_FOR;
   #commands := #clear_commands;
   #commands.out.done := TRUE;
END_FUNCTION

// folder: OBs

ORGANIZATION_BLOCK "Rack or station failure"   // OB86, LAD, RackStationFailure
{ S7_Optimized_Access := 'TRUE' }
VERSION : 0.1
   VAR_INPUT
      LADDR : Hw_Device;   // Hardware identifier
      Event_Class : Byte;   // Event class
      Fault_ID : Byte;   // Fault identifier
   END_VAR
BEGIN
END_ORGANIZATION_BLOCK

ORGANIZATION_BLOCK "Startup"   // OB100, LAD, Startup
TITLE = "Complete Restart"
{ S7_Optimized_Access := 'TRUE' }
VERSION : 0.1
   VAR_INPUT
      LostRetentive : Bool;   // True if retentive data are lost
      LostRTC : Bool;   // True if date and time are lost
   END_VAR
BEGIN

REGION Network 1 (SCL): HMI STATION INITIALIZATION
END_REGION
END_ORGANIZATION_BLOCK

ORGANIZATION_BLOCK "Programming error"   // OB121, LAD, ProgrammingError
{ S7_Optimized_Access := 'TRUE' }
VERSION : 0.1
   VAR_INPUT
      BlockNr : UInt;   // Number of causing block
      Reaction : USInt;   // 0:ignore, 1:substitute, 2:skip
      Fault_ID : Byte;   // Fault identifier
      BlockType : USInt;   // 16#01:OB, 16#02:FC, 16#03:FB, 16#04:SFC, 16#05:SFB, 16#06:DB: Type of block causing the error
      Area : USInt;   // Area where the error occured
      DBNr : DB_ANY;   // DB number if Area = DB or DI
      Csg_OBNr : OB_Any;   // Number of OB causing the error
      Csg_Prio : USInt;   // Priority of OB causing the error
      Width : USInt;   // 0:bit, 1:byte, 2:word, 3:dword, 4:lword
   END_VAR
BEGIN
END_ORGANIZATION_BLOCK

ORGANIZATION_BLOCK "IO access error"   // OB122, LAD, IOAccessError
{ S7_Optimized_Access := 'TRUE' }
VERSION : 0.1
   VAR_INPUT
      BlockNr : UInt;   // Number of causing block
      Reaction : USInt;   // 0:ignore, 1:substitute, 2:skip
      Fault_ID : Byte;   // 16#42:reading, 16#43:writing
      BlockType : USInt;   // 16#01:OB, 16#02:FC, 16#03:FB, 16#04:SFC, 16#05:SFB, 16#06:DB: Type of block causing the error
      Area : USInt;   // 16#81:I, 16#82:Q: IO area where the IOaccess error occured
      DBNr : DB_ANY;   // Reserved for system
      Csg_OBNr : OB_Any;   // Number of OB causing the error
      Csg_Prio : USInt;   // Priority of OB causing the error
      Width : USInt;   // 0:bit, 1:byte, 2:word, 3:dword, 4:lword
   END_VAR
BEGIN
END_ORGANIZATION_BLOCK

// folder: Order/States

FUNCTION_BLOCK "Order State"   // FB2, SCL
{ S7_Optimized_Access := 'TRUE' }
VERSION : 0.1
   VAR_INPUT
      pnLib : "Recipe: PN Text Library";
   END_VAR
   VAR_IN_OUT
      stns : "Station: All Stations";
   END_VAR
   VAR_TEMP
      pStn : Int;
      pBtn : Int;
      stn : "Station: Single Station";
   END_VAR
BEGIN
   REGION "FOR EACH STATION"
       FOR #pStn := 0 TO "STATION_COUNT" DO

           REGION "FOR EACH BUTTON"
               FOR #pBtn := 0 TO "STATION_BUTTON_COUNT" DO

                   REGION "POPULATE CURRENT STATION"
                       #stn := #stns.stn[#pStn];
                   END_REGION

                   REGION "INITIALIZE STATE"
                       "Order State: Initialize State"(newParams := #stn.wipCmpts.flags.newPN,
                                                       pnGood := #stn.wipCmpts.flags.pnGood[#pBtn],
                                                       state := #stn.wipCmpts.orderState[#pBtn]);
                   END_REGION

                   REGION "ENTER IDLE"
                       "Order State: Enter Idle"(btnFalling := #stn.wipCmpts.kp8Logical.falling.btn[#pBtn],
                                                 state := #stn.wipCmpts.orderState[#pBtn]);
                   END_REGION

                   REGION "ENTER REQUESTED"
                       "Order State: Enter Requested"(btnRising := #stn.wipCmpts.kp8Logical.rising.btn[#pBtn],
                                                      state := #stn.wipCmpts.orderState[#pBtn]);
                   END_REGION

                   REGION "ENTER REQUESTED CRITICAL"
                       "Order State: Enter Requested Critical"(timerVal := #stn.wipCmpts.timers.remaining[#pBtn],
                                                               state := #stn.wipCmpts.orderState[#pBtn]);
                   END_REGION

                   REGION "ENTER REQUESTED EXPIRED"
                       "Order State: Enter Requested Expired"(timerVal := #stn.wipCmpts.timers.remaining[#pBtn],
                                                              state := #stn.wipCmpts.orderState[#pBtn]);
                   END_REGION

                   REGION "SAVE CURRENT STATION"
                       #stns.stn[#pStn] := #stn;
                   END_REGION

               END_FOR;
           END_REGION

       END_FOR;
   END_REGION
END_FUNCTION_BLOCK

FUNCTION "Order State: Enter Idle" : Void   // FC6, SCL
{ S7_Optimized_Access := 'TRUE' }
VERSION : 0.1
   VAR_INPUT
      btnFalling : Bool;
   END_VAR
   VAR_IN_OUT
      state : Int;
   END_VAR
BEGIN
   IF #btnFalling THEN
       #state := "idle";
   END_IF;
END_FUNCTION

FUNCTION "Order State: Enter Requested" : Void   // FC7, SCL
{ S7_Optimized_Access := 'TRUE' }
VERSION : 0.1
   VAR_INPUT
      btnRising : Bool;
   END_VAR
   VAR_IN_OUT
      state : Int;
   END_VAR
BEGIN
   IF #state = "idle" THEN
       IF #btnRising THEN
           #state := "requested";
       END_IF;
   END_IF;
END_FUNCTION

FUNCTION "Order State: Initialize State" : Void   // FC10, SCL
{ S7_Optimized_Access := 'TRUE' }
VERSION : 0.1
   VAR_INPUT
      newParams : Bool;
      pnGood : Bool;
   END_VAR
   VAR_IN_OUT
      state : Int;
   END_VAR
BEGIN
   REGION "ON NEW PARAMETERS"
       IF #newParams THEN

           REGION "ON VALID PN" 
               IF #pnGood THEN

                   REGION "INITIALIZE STATE"
                       #state := BOOL_TO_INT(#pnGood);
                   END_REGION